        [210].Name := 'Mary', [210].Class := 'Foundation', [211].Name := 'Mary', [211].Class := 'Registered', [212].Name := 'Northwest Tandem', [212].Class := 'Certified', [213].Name := 'Northwest Tandem', [213].Class := 'Common', [214].Name := 'Northwest Tandem', [214].Class := 'Foundation', [215].Name := 'Northwest Tandem', [215].Class := 'Registered', [216].Name := 'NW Duet', [216].Class := 'Certified', [217].Name := 'NW Duet', [217].Class := 'Common', [218].Name := 'NW Duet', [218].Class := 'Foundation', [219].Name := 'NW Duet', [219].Class := 'Registered', [220].Name := 'ORCF 101', [220].Class := 'Certified', [221].Name := 'ORCF 101', [221].Class := 'Common', [222].Name := 'ORCF 101', [222].Class := 'Foundation', [223].Name := 'ORCF 101', [223].Class := 'Registered', [224].Name := 'ORCF 102', [224].Class := 'Certified', [225].Name := 'ORCF 102', [225].Class := 'Common', [226].Name := 'ORCF 102', [226].Class := 'Foundation', [227].Name := 'ORCF 102', [227].Class := 'Registered', [228].Name := 'Ovation', [228].Class := 'Certified', [229].Name := 'Ovation', [229].Class := 'Common', [230].Name := 'Ovation', [230].Class := 'Foundation', [231].Name := 'Ovation', [231].Class := 'Registered', [232].Name := 'Palouse', [232].Class := 'Certified', [233].Name := 'Palouse', [233].Class := 'Common', [234].Name := 'Palouse', [234].Class := 'Foundation', [235].Name := 'Palouse', [235].Class := 'Registered', [236].Name := 'Puma', [236].Class := 'Certified', [237].Name := 'Puma', [237].Class := 'Common', [238].Name := 'Puma', [238].Class := 'Foundation', [239].Name := 'Puma', [239].Class := 'Registered',
        [240].Name := 'Rod', [240].Class := 'Certified', [241].Name := 'Rod', [241].Class := 'Common', [242].Name := 'Rod', [242].Class := 'Foundation', [243].Name := 'Rod', [243].Class := 'Registered', [244].Name := 'Scotch-Spokane Seed', [244].Class := 'Certified', [245].Name := 'Scotch-Spokane Seed', [245].Class := 'Common', [246].Name := 'Scotch-Spokane Seed', [246].Class := 'Foundation', [247].Name := 'Scotch-Spokane Seed', [247].Class := 'Registered', [248].Name := 'Scotch-Spokane Seed-Day', [248].Class := 'Certified', [249].Name := 'Scotch-Spokane Seed-Day', [249].Class := 'Common', [250].Name := 'Scotch-Spokane Seed-Day', [250].Class := 'Foundation', [251].Name := 'Scotch-Spokane Seed-Day', [251].Class := 'Registered', [252].Name := 'Seahawk', [252].Class := 'Certified', [253].Name := 'Seahawk', [253].Class := 'Common', [254].Name := 'Seahawk', [254].Class := 'Foundation', [255].Name := 'Seahawk', [255].Class := 'Registered', [256].Name := 'Sierra', [256].Class := 'Certified', [257].Name := 'Sierra', [257].Class := 'Common', [258].Name := 'Sierra', [258].Class := 'Foundation', [259].Name := 'Sierra', [259].Class := 'Registered', [260].Name := 'Sierra PNWFC', [260].Class := 'Certified', [261].Name := 'Sierra PNWFC', [261].Class := 'Common', [262].Name := 'Sierra PNWFC', [262].Class := 'Foundation', [263].Name := 'Sierra PNWFC', [263].Class := 'Registered', [264].Name := 'Sierra Spokane Seed', [264].Class := 'Certified', [265].Name := 'Sierra Spokane Seed', [265].Class := 'Common', [266].Name := 'Sierra Spokane Seed', [266].Class := 'Foundation', [267].Name := 'Sierra Spokane Seed', [267].Class := 'Registered', [268].Name := 'Skiles', [268].Class := 'Certified', [269].Name := 'Skiles', [269].Class := 'Common',
        [270].Name := 'Skiles', [270].Class := 'Foundation', [271].Name := 'Skiles', [271].Class := 'Registered', [272].Name := 'Solano', [272].Class := 'Certified', [273].Name := 'Solano', [273].Class := 'Common', [274].Name := 'Solano', [274].Class := 'Foundation', [275].Name := 'Solano', [275].Class := 'Registered', [276].Name := 'Stephens', [276].Class := 'Certified', [277].Name := 'Stephens', [277].Class := 'Common', [278].Name := 'Stephens', [278].Class := 'Foundation', [279].Name := 'Stephens', [279].Class := 'Registered', [280].Name := 'Sy 107', [280].Class := 'Certified', [281].Name := 'Sy 107', [281].Class := 'Common', [282].Name := 'Sy 107', [282].Class := 'Foundation', [283].Name := 'Sy 107', [283].Class := 'Registered', [284].Name := 'SY 605', [284].Class := 'Certified', [285].Name := 'SY 605', [285].Class := 'Common', [286].Name := 'SY 605', [286].Class := 'Foundation', [287].Name := 'SY 605', [287].Class := 'Registered', [288].Name := 'SY Assure', [288].Class := 'Certified', [289].Name := 'SY Assure', [289].Class := 'Common', [290].Name := 'SY Assure', [290].Class := 'Foundation', [291].Name := 'SY Assure', [291].Class := 'Registered', [292].Name := 'Test', [292].Class := 'Certified', [293].Name := 'Test', [293].Class := 'Common', [294].Name := 'Test', [294].Class := 'Foundation', [295].Name := 'Test', [295].Class := 'Registered', [296].Name := 'Tubbs', [296].Class := 'Certified', [297].Name := 'Tubbs', [297].Class := 'Common', [298].Name := 'Tubbs', [298].Class := 'Foundation', [299].Name := 'Tubbs', [299].Class := 'Registered',
        [300].Name := 'Universal-Spokane Seed', [300].Class := 'Certified', [301].Name := 'Universal-Spokane Seed', [301].Class := 'Common', [302].Name := 'Universal-Spokane Seed', [302].Class := 'Foundation', [303].Name := 'Universal-Spokane Seed', [303].Class := 'Registered', [304].Name := 'Vespa', [304].Class := 'Certified', [305].Name := 'Vespa', [305].Class := 'Common', [306].Name := 'Vespa', [306].Class := 'Foundation', [307].Name := 'Vespa', [307].Class := 'Registered', [308].Name := 'WB 1035 CL spring', [308].Class := 'Certified', [309].Name := 'WB 1035 CL spring', [309].Class := 'Common', [310].Name := 'WB 1035 CL spring', [310].Class := 'Foundation', [311].Name := 'WB 1035 CL spring', [311].Class := 'Registered', [312].Name := 'WB 1070', [312].Class := 'Certified', [313].Name := 'WB 1070', [313].Class := 'Common', [314].Name := 'WB 1070', [314].Class := 'Foundation', [315].Name := 'WB 1070', [315].Class := 'Registered', [316].Name := 'WB 1376', [316].Class := 'Certified', [317].Name := 'WB 1376', [317].Class := 'Common', [318].Name := 'WB 1376', [318].Class := 'Foundation', [319].Name := 'WB 1376', [319].Class := 'Registered', [320].Name := 'WB 1529', [320].Class := 'Certified', [321].Name := 'WB 1529', [321].Class := 'Common', [322].Name := 'WB 1529', [322].Class := 'Foundation', [323].Name := 'WB 1529', [323].Class := 'Registered', [324].Name := 'WB 1604', [324].Class := 'Certified', [325].Name := 'WB 1604', [325].Class := 'Common', [326].Name := 'WB 1604', [326].Class := 'Foundation', [327].Name := 'WB 1604', [327].Class := 'Registered', [328].Name := 'WB 528', [328].Class := 'Certified', [329].Name := 'WB 528', [329].Class := 'Common',
        [330].Name := 'WB 528', [330].Class := 'Foundation', [331].Name := 'WB 528', [331].Class := 'Registered', [332].Name := 'WB 6121 spring', [332].Class := 'Certified', [333].Name := 'WB 6121 spring', [333].Class := 'Common', [334].Name := 'WB 6121 spring', [334].Class := 'Foundation', [335].Name := 'WB 6121 spring', [335].Class := 'Registered', [336].Name := 'WB 6341 Spring', [336].Class := 'Certified', [337].Name := 'WB 6341 Spring', [337].Class := 'Common', [338].Name := 'WB 6341 Spring', [338].Class := 'Foundation', [339].Name := 'WB 6341 Spring', [339].Class := 'Registered', [340].Name := 'WB 9411', [340].Class := 'Certified', [341].Name := 'WB 9411', [341].Class := 'Common', [342].Name := 'WB 9411', [342].Class := 'Foundation', [343].Name := 'WB 9411', [343].Class := 'Registered', [344].Name := 'WB 9518', [344].Class := 'Certified', [345].Name := 'WB 9518', [345].Class := 'Common', [346].Name := 'WB 9518', [346].Class := 'Foundation', [347].Name := 'WB 9518', [347].Class := 'Registered', [348].Name := 'WB523', [348].Class := 'Certified', [349].Name := 'WB523', [349].Class := 'Common', [350].Name := 'WB523', [350].Class := 'Foundation', [351].Name := 'WB523', [351].Class := 'Registered', [352].Name := 'Xerpha', [352].Class := 'Certified', [353].Name := 'Xerpha', [353].Class := 'Common', [354].Name := 'Xerpha', [354].Class := 'Foundation', [355].Name := 'Xerpha', [355].Class := 'Registered');
   varIndx : DINT;
   vartableONS : DINT := 3;
   VarTrimTemp : STRING := '843001';
   VIRTUAL_BT : ALIAS FOR N20[5].13;
   VIRTUAL_BT1 : ALIAS FOR N23[0].12;
   VIRTUAL_BT2 : ALIAS FOR N23[0].13;
   zzzRealtmp : REAL := 30.73328;
   zzzsqlVaritiesRevd : BOOL;
   zzztmpSqlDataArryDINT : DINT[10];
   zzztmpSqlDataArryFLT : REAL[10];
   zzztmpSqlDataDINT : DINT := 1000;
   zzztmpSqlDataFLT : REAL;
   zzztmpSqlDataSTR : STRING;
   zzztmpTANKtest : DINT[10];
   zzzz_22_GATE_PO_STOR : DINT;
   zzzzProcessAll : DINT;
   zzzzSTRING : STRING := '821001 ArtDeco SWW';
   zzzzTestGrossWt : BOOL;
   zzzzTestTareWt : BOOL;
   zzzztmpDINT : DINT[10];
   zzzzVAR_CNT_ONS : BOOL;
   zzzzzTestBit : BOOL;
END_VAR

PROGRAM _2_MAIN   (* main routine _02_MAIN *)
VAR
   Flow_Gal2Oz : FBD_MATH := (SourceB := 0.015);
   GRT_01 : FBD_COMPARE := (SourceB := 75.0);
   HOUR_METERS : DINT;
   LES_01 : FBD_COMPARE;
   LES_02 : FBD_COMPARE;
   SCL_01 : SCALE := (InRawMax := 100.0, InEUMax := 4000.0);
   SCL_02 : SCALE := (In := 28776.0, InRawMin := 31000.0, InEUMax := 3200.0, Status := 16#0000_0003, InstructFault := 1, InRawRangeInv := 1);
   SCL_03 : SCALE := (In := 6569.0, InRawMax := 13975.0, InRawMin := 578.0, InEUMax := 3000.0, Out := 1341.569);
   SCL_04 : SCALE;
   SCL_05 : SCALE;
   SCL_06 : SCALE := (InRawMax := 60.0, InEUMax := 32767.0);
   SCL_07 : SCALE := (In := 46.0, InRawMax := 60.0, InEUMax := 31000.0, Out := 23766.668);
   SCL_08 : SCALE := (In := 48.0, InRawMax := 60.0, InEUMax := 31000.0, Out := 24800.0);
   SCL_09 : SCALE := (In := 53.0, InRawMax := 60.0, InEUMax := 31000.0, Out := 27383.334);
   SEL_01 : SELECT;
   SUB_01 : FBD_MATH;
   Test_Bit : BOOL;
   TOT_01 : TOTALIZER := (Gain := 1.0, ProgProgReq := 1, ProgStartReq := 1, RTSTime := 1, Total := 3307.86, OldTotal := 877.80005, ProgOper := 1, RunStop := 1, TargetFlag := 1, TargetDev1Flag := 1, TargetDev2Flag := 1, LowInCutoffFlag := 1, DeltaT := 0.004);
END_VAR

ROUTINE _02_MAIN   (* ladder *)
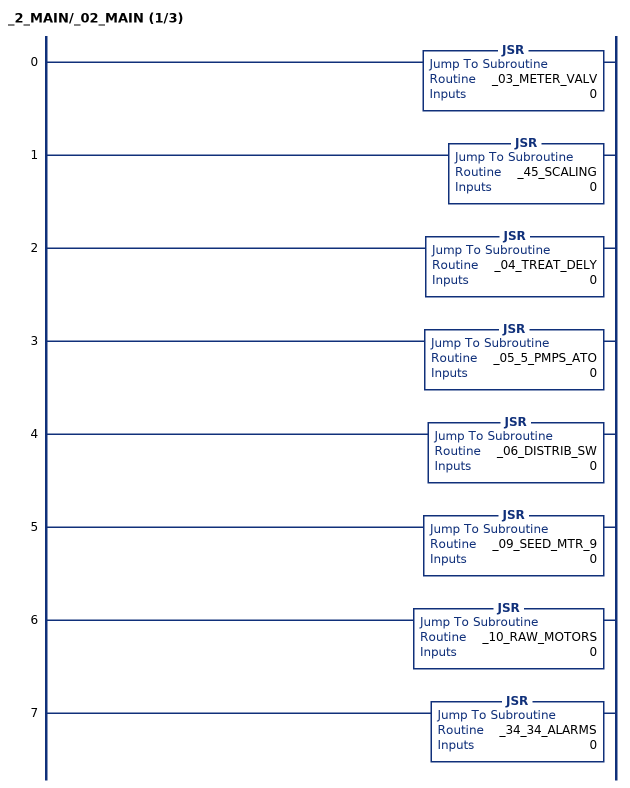
   0: JSR(_03_METER_VALV,0);
   1: JSR(_45_SCALING,0);
   2: JSR(_04_TREAT_DELY,0);
   3: JSR(_05_5_PMPS_ATO,0);
   4: JSR(_06_DISTRIB_SW,0);
   5: JSR(_09_SEED_MTR_9,0);
   6: JSR(_10_RAW_MOTORS,0);
   7: JSR(_34_34_ALARMS,0);
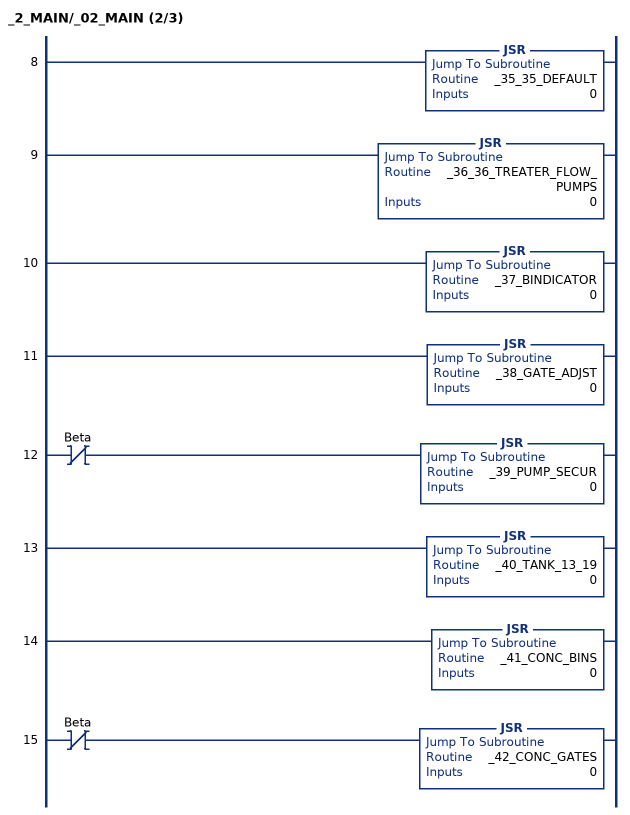
   8: JSR(_35_35_DEFAULT,0);
   9: JSR(_36_36_TREATER_FLOW_PUMPS,0);
   10: JSR(_37_BINDICATOR,0);
   11: JSR(_38_GATE_ADJST,0);
   12: XIO(Beta)JSR(_39_PUMP_SECUR,0);
   13: JSR(_40_TANK_13_19,0);
   14: JSR(_41_CONC_BINS,0);
   15: XIO(Beta)JSR(_42_CONC_GATES,0);
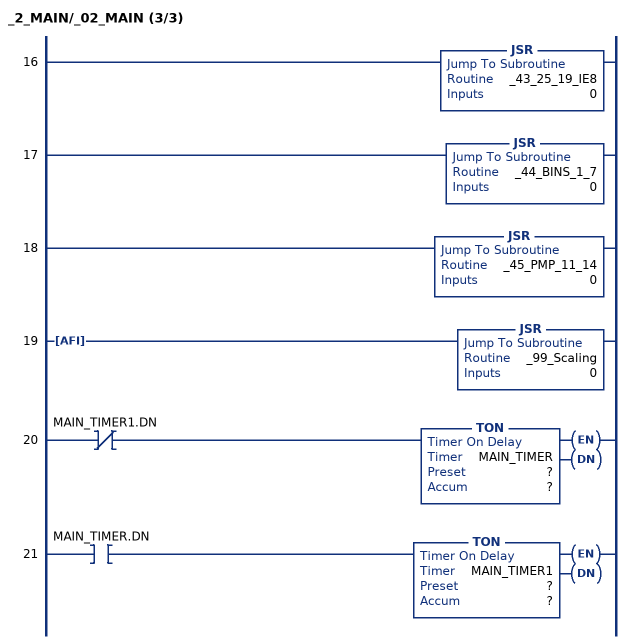
   16: JSR(_43_25_19_IE8,0);
   17: JSR(_44_BINS_1_7,0);
   18: JSR(_45_PMP_11_14,0);
   19: AFI()JSR(_99_Scaling,0);
   20: XIO(MAIN_TIMER1.DN)TON(MAIN_TIMER,?,?);
   21: XIC(MAIN_TIMER.DN)TON(MAIN_TIMER1,?,?);
END_ROUTINE

ROUTINE _03_METER_VALV   (* ladder *)
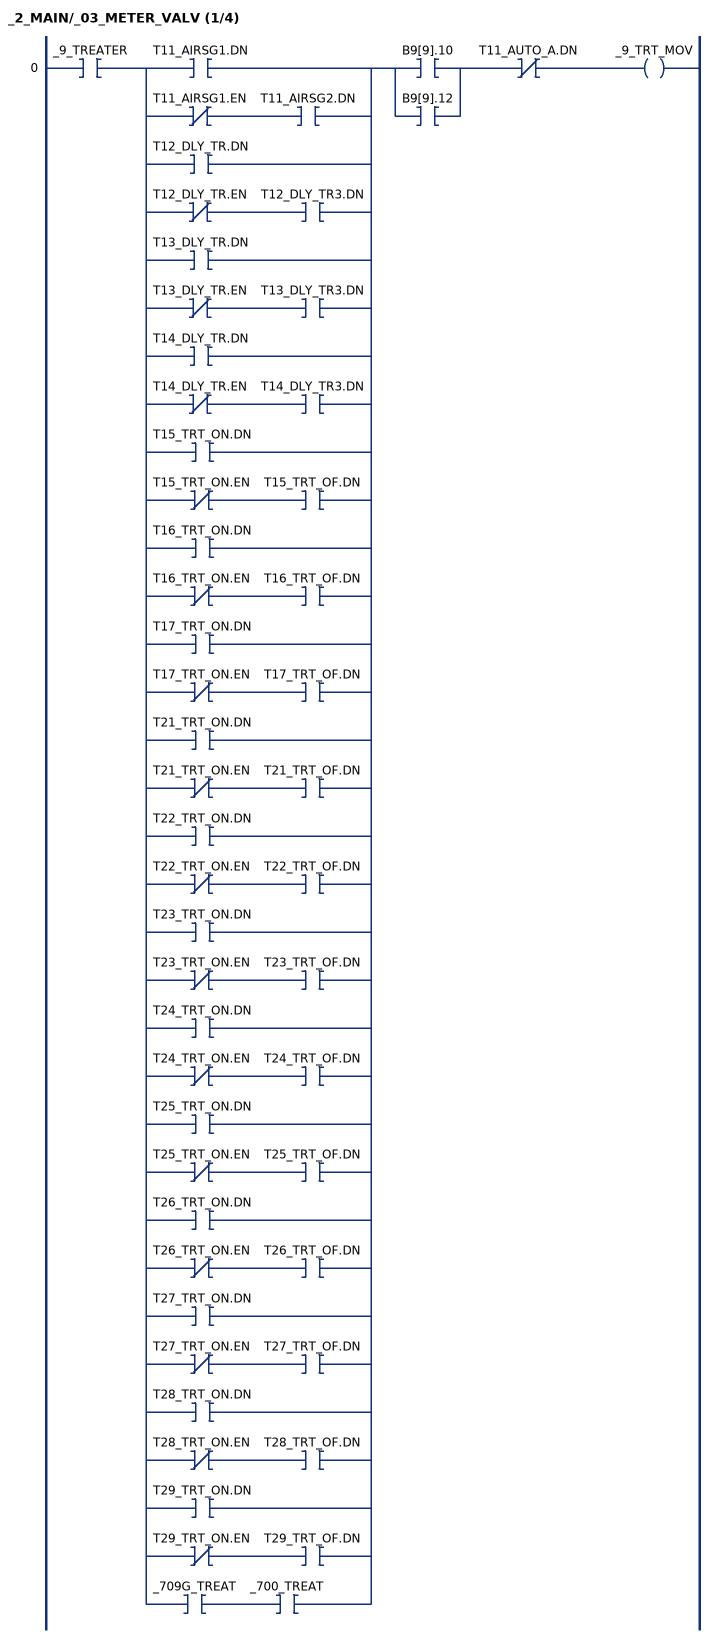
   0: XIC(_9_TREATER)[XIC(T11_AIRSG1.DN) ,XIO(T11_AIRSG1.EN) XIC(T11_AIRSG2.DN) ,XIC(T12_DLY_TR.DN) ,XIO(T12_DLY_TR.EN) XIC(T12_DLY_TR3.DN) ,XIC(T13_DLY_TR.DN) ,XIO(T13_DLY_TR.EN) XIC(T13_DLY_TR3.DN) ,XIC(T14_DLY_TR.DN) ,XIO(T14_DLY_TR.EN) XIC(T14_DLY_TR3.DN) ,XIC(T15_TRT_ON.DN) ,XIO(T15_TRT_ON.EN) XIC(T15_TRT_OF.DN) ,XIC(T16_TRT_ON.DN) ,XIO(T16_TRT_ON.EN) XIC(T16_TRT_OF.DN) ,XIC(T17_TRT_ON.DN) ,XIO(T17_TRT_ON.EN) XIC(T17_TRT_OF.DN) ,XIC(T21_TRT_ON.DN) ,XIO(T21_TRT_ON.EN) XIC(T21_TRT_OF.DN) ,XIC(T22_TRT_ON.DN) ,XIO(T22_TRT_ON.EN) XIC(T22_TRT_OF.DN) ,XIC(T23_TRT_ON.DN) ,XIO(T23_TRT_ON.EN) XIC(T23_TRT_OF.DN) ,XIC(T24_TRT_ON.DN) ,XIO(T24_TRT_ON.EN) XIC(T24_TRT_OF.DN) ,XIC(T25_TRT_ON.DN) ,XIO(T25_TRT_ON.EN) XIC(T25_TRT_OF.DN) ,XIC(T26_TRT_ON.DN) ,XIO(T26_TRT_ON.EN) XIC(T26_TRT_OF.DN) ,XIC(T27_TRT_ON.DN) ,XIO(T27_TRT_ON.EN) XIC(T27_TRT_OF.DN) ,XIC(T28_TRT_ON.DN) ,XIO(T28_TRT_ON.EN) XIC(T28_TRT_OF.DN) ,XIC(T29_TRT_ON.DN) ,XIO(T29_TRT_ON.EN) XIC(T29_TRT_OF.DN) ,XIC(_709G_TREAT) XIC(_700_TREAT) ][XIC(B9[9].10) ,XIC(B9[9].12) ]XIO(T11_AUTO_A.DN)OTE(_9_TRT_MOV);
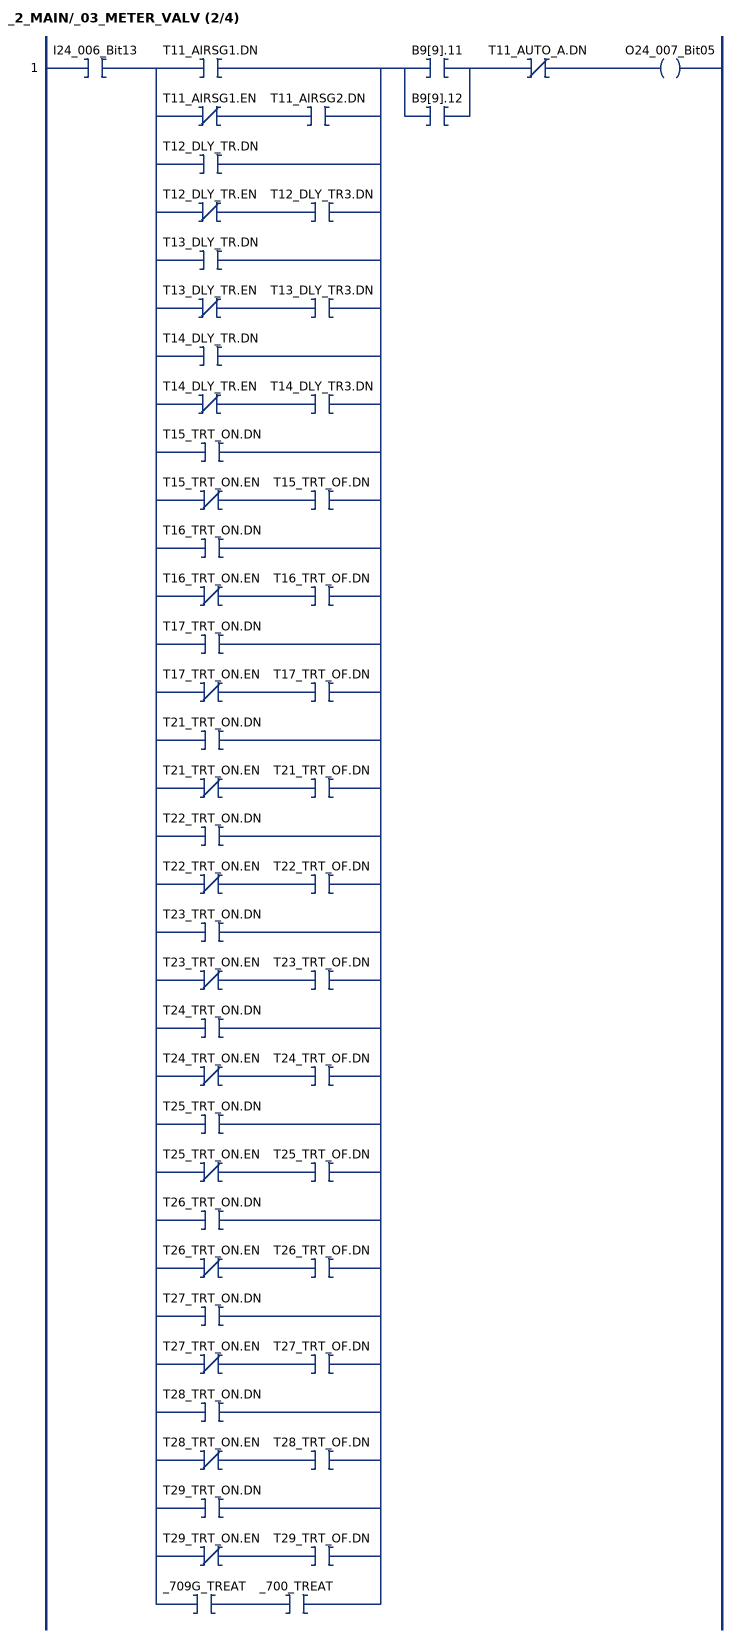
   1: XIC(I24_006_Bit13)[XIC(T11_AIRSG1.DN) ,XIO(T11_AIRSG1.EN) XIC(T11_AIRSG2.DN) ,XIC(T12_DLY_TR.DN) ,XIO(T12_DLY_TR.EN) XIC(T12_DLY_TR3.DN) ,XIC(T13_DLY_TR.DN) ,XIO(T13_DLY_TR.EN) XIC(T13_DLY_TR3.DN) ,XIC(T14_DLY_TR.DN) ,XIO(T14_DLY_TR.EN) XIC(T14_DLY_TR3.DN) ,XIC(T15_TRT_ON.DN) ,XIO(T15_TRT_ON.EN) XIC(T15_TRT_OF.DN) ,XIC(T16_TRT_ON.DN) ,XIO(T16_TRT_ON.EN) XIC(T16_TRT_OF.DN) ,XIC(T17_TRT_ON.DN) ,XIO(T17_TRT_ON.EN) XIC(T17_TRT_OF.DN) ,XIC(T21_TRT_ON.DN) ,XIO(T21_TRT_ON.EN) XIC(T21_TRT_OF.DN) ,XIC(T22_TRT_ON.DN) ,XIO(T22_TRT_ON.EN) XIC(T22_TRT_OF.DN) ,XIC(T23_TRT_ON.DN) ,XIO(T23_TRT_ON.EN) XIC(T23_TRT_OF.DN) ,XIC(T24_TRT_ON.DN) ,XIO(T24_TRT_ON.EN) XIC(T24_TRT_OF.DN) ,XIC(T25_TRT_ON.DN) ,XIO(T25_TRT_ON.EN) XIC(T25_TRT_OF.DN) ,XIC(T26_TRT_ON.DN) ,XIO(T26_TRT_ON.EN) XIC(T26_TRT_OF.DN) ,XIC(T27_TRT_ON.DN) ,XIO(T27_TRT_ON.EN) XIC(T27_TRT_OF.DN) ,XIC(T28_TRT_ON.DN) ,XIO(T28_TRT_ON.EN) XIC(T28_TRT_OF.DN) ,XIC(T29_TRT_ON.DN) ,XIO(T29_TRT_ON.EN) XIC(T29_TRT_OF.DN) ,XIC(_709G_TREAT) XIC(_700_TREAT) ][XIC(B9[9].11) ,XIC(B9[9].12) ]XIO(T11_AUTO_A.DN)OTE(O24_007_Bit05);
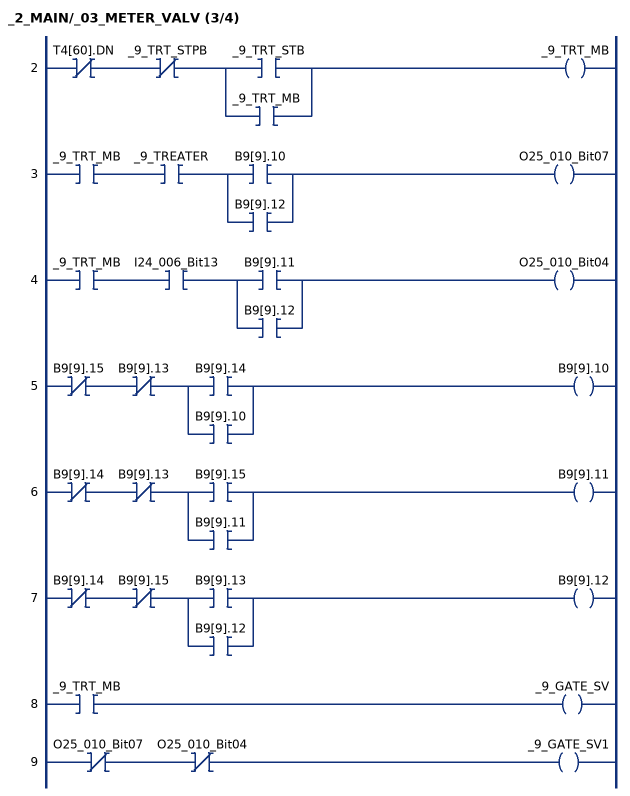
   2: XIO(T4[60].DN)XIO(_9_TRT_STPB)[XIC(_9_TRT_STB) ,XIC(_9_TRT_MB) ]OTE(_9_TRT_MB);
   3: XIC(_9_TRT_MB)XIC(_9_TREATER)[XIC(B9[9].10) ,XIC(B9[9].12) ]OTE(O25_010_Bit07);
   4: XIC(_9_TRT_MB)XIC(I24_006_Bit13)[XIC(B9[9].11) ,XIC(B9[9].12) ]OTE(O25_010_Bit04);
   5: XIO(B9[9].15)XIO(B9[9].13)[XIC(B9[9].14) ,XIC(B9[9].10) ]OTE(B9[9].10);
   6: XIO(B9[9].14)XIO(B9[9].13)[XIC(B9[9].15) ,XIC(B9[9].11) ]OTE(B9[9].11);
   7: XIO(B9[9].14)XIO(B9[9].15)[XIC(B9[9].13) ,XIC(B9[9].12) ]OTE(B9[9].12);
   8: XIC(_9_TRT_MB)OTE(_9_GATE_SV);
   9: XIO(O25_010_Bit07)XIO(O25_010_Bit04)OTE(_9_GATE_SV1);